VERSION : 0.1
   VAR
      ReadWriteDeviceNo : Int := 0;
      CopyDeviceNO : Int := 0;
      Read : Bool := FALSE;
      Write : Bool := FALSE;
      Copy : Bool := FALSE;
      Option : Array[0..2] of Struct
         With2PSwitch : Bool;
      END_STRUCT;
      MH_Hyd : Array[0..2] of "UDT721_Hydraulic";
      S_Hyd : Array[0..2] of "UDT721_Hydraulic";
      NZL_Hyd : Array[0..2] of "UDT721_Hydraulic";
   END_VAR
BEGIN
   MH_Hyd[0].Hyd_Filter_supervision := S5T#30S;
   MH_Hyd[0].Hyd_P_Startup := S5T#15S;
   MH_Hyd[0].Hyd_P_Supervision := S5T#5S;
   MH_Hyd[0].Hyd_CP_Time := S5T#4S;
   MH_Hyd[0].Hyd_PressureSwitch := S5T#0MS;
   MH_Hyd[0].Hyd_SwitchOFFDelay := S5T#0MS;
   MH_Hyd[1].Hyd_Filter_supervision := S5T#30S;
   MH_Hyd[1].Hyd_P_Startup := S5T#15S;
   MH_Hyd[1].Hyd_P_Supervision := S5T#5S;
   MH_Hyd[1].Hyd_CP_Time := S5T#4S;
   MH_Hyd[1].Hyd_PressureSwitch := S5T#0MS;
   MH_Hyd[1].Hyd_SwitchOFFDelay := S5T#0MS;
   MH_Hyd[2].Hyd_Filter_supervision := S5T#0MS;
   MH_Hyd[2].Hyd_P_Startup := S5T#0MS;
   MH_Hyd[2].Hyd_P_Supervision := S5T#0MS;
   MH_Hyd[2].Hyd_CP_Time := S5T#0MS;
   MH_Hyd[2].Hyd_PressureSwitch := S5T#0MS;
   MH_Hyd[2].Hyd_SwitchOFFDelay := S5T#0MS;
   S_Hyd[0].Hyd_Filter_supervision := S5T#0MS;
   S_Hyd[0].Hyd_P_Startup := S5T#0MS;
   S_Hyd[0].Hyd_P_Supervision := S5T#0MS;
   S_Hyd[0].Hyd_CP_Time := S5T#0MS;
   S_Hyd[0].Hyd_PressureSwitch := S5T#0MS;
   S_Hyd[0].Hyd_SwitchOFFDelay := S5T#0MS;
   S_Hyd[1].Hyd_Filter_supervision := S5T#0MS;
   S_Hyd[1].Hyd_P_Startup := S5T#0MS;
   S_Hyd[1].Hyd_P_Supervision := S5T#0MS;
   S_Hyd[1].Hyd_CP_Time := S5T#0MS;
   S_Hyd[1].Hyd_PressureSwitch := S5T#0MS;
   S_Hyd[1].Hyd_SwitchOFFDelay := S5T#0MS;
   S_Hyd[2].Hyd_Filter_supervision := S5T#0MS;
   S_Hyd[2].Hyd_P_Startup := S5T#0MS;
   S_Hyd[2].Hyd_P_Supervision := S5T#0MS;
   S_Hyd[2].Hyd_CP_Time := S5T#0MS;
   S_Hyd[2].Hyd_PressureSwitch := S5T#0MS;
   S_Hyd[2].Hyd_SwitchOFFDelay := S5T#0MS;
   NZL_Hyd[0].Hyd_Filter_supervision := S5T#0MS;
   NZL_Hyd[0].Hyd_P_Startup := S5T#0MS;
   NZL_Hyd[0].Hyd_P_Supervision := S5T#0MS;
   NZL_Hyd[0].Hyd_CP_Time := S5T#0MS;
   NZL_Hyd[0].Hyd_PressureSwitch := S5T#0MS;
   NZL_Hyd[0].Hyd_SwitchOFFDelay := S5T#0MS;
   NZL_Hyd[1].Hyd_Filter_supervision := S5T#0MS;
   NZL_Hyd[1].Hyd_P_Startup := S5T#0MS;
   NZL_Hyd[1].Hyd_P_Supervision := S5T#0MS;
   NZL_Hyd[1].Hyd_CP_Time := S5T#0MS;
   NZL_Hyd[1].Hyd_PressureSwitch := S5T#0MS;
   NZL_Hyd[1].Hyd_SwitchOFFDelay := S5T#0MS;
   NZL_Hyd[2].Hyd_Filter_supervision := S5T#0MS;
   NZL_Hyd[2].Hyd_P_Startup := S5T#0MS;
   NZL_Hyd[2].Hyd_P_Supervision := S5T#0MS;
   NZL_Hyd[2].Hyd_CP_Time := S5T#0MS;
   NZL_Hyd[2].Hyd_PressureSwitch := S5T#0MS;
   NZL_Hyd[2].Hyd_SwitchOFFDelay := S5T#0MS;
   Option[0].With2PSwitch := TRUE;
   Option[1].With2PSwitch := TRUE;
   Option[2].With2PSwitch := FALSE;
END_DATA_BLOCK

DATA_BLOCK "DB753_MeteringPump"   // DB753
TITLE = Parameter metering pump
{ S7_Optimized_Access := 'FALSE' }
NAME : metering
VERSION : 0.1
   VAR
      ReadWriteDeviceNo : Int := 0;
      CopyDeviceNO : Int := 0;
      Read : Bool := FALSE;
      Write : Bool := FALSE;
      Copy : Bool := FALSE;
      Pump : Array[0..12] of "UDT753_MeteringPump";
      Heating : Array[0..12] of Struct
         Exist : Array[1..8] of Bool;
      END_STRUCT;
      HeatingController : Array[0..4] of Struct
         Heating : Array[1..8] of "UDT702_HeatingControl";
      END_STRUCT;
   END_VAR
BEGIN
   Pump[0].Pump_Active := TRUE;
   Pump[0].WithFC := TRUE;
   Pump[0].WithoutFlowControl := TRUE;
   Pump[0].WithFeedPump := FALSE;
   Pump[0].WithEdgeFilter := FALSE;
   Pump[0].MachineNumber := 16#01;
   Pump[0]."Name" := 'Poly';
   Pump[0].TankNo := 1;
   Pump[0].Pulse_per_liter := 333.333;
   Pump[1].Pump_Active := TRUE;
   Pump[1].WithFC := TRUE;
   Pump[1].WithoutFlowControl := TRUE;
   Pump[1].WithFeedPump := FALSE;
   Pump[1].WithEdgeFilter := FALSE;
   Pump[1]."Name" := 'Poly';
   Pump[1].TankNo := 1;
   Pump[2].Pump_Active := TRUE;
   Pump[2].WithFC := TRUE;
   Pump[2].WithoutFlowControl := TRUE;
   Pump[2].WithFeedPump := FALSE;
   Pump[2].WithEdgeFilter := FALSE;
   Pump[2].MachineNumber := 16#01;
   Pump[2]."Name" := 'Iso';
   Pump[2].TankNo := 2;
   Pump[2].Pulse_per_liter := 965.667;
   Pump[0].Flow_State := 16#0000;
   Pump[0].RunTimePumpInterval := S5T#0MS;
   Pump[0].PauseTimePumpInterval := S5T#0MS;
   Pump[0].Flow_Index := 16#0000;
   Pump[0].DelayPressureFeedP := S5T#9S;
   Pump[0].DelayRunTimeFeedP := S5T#6S;
   Pump[0].MinTempRelease := 0.0;
   Pump[0].With_2Point := FALSE;
   Pump[0].WithFlowControl := FALSE;
   Pump[0].PumDeselectionEnable := FALSE;
   Pump[0].PumpDeselected := FALSE;
   Pump[0].PumpDeselectedInterval := FALSE;
   Pump[0].WithFischerValveHP := FALSE;
   Pump[0].WithFischerValveLP := FALSE;
   Pump[0].WithHPHeatExchanger := FALSE;
   Pump[0].WithLPHeatExchanger := FALSE;
   Pump[0].WithExhauseSystem := FALSE;
   Pump[0].WithHeating := FALSE;
   Pump[0].WithPipeHeating := FALSE;
   Pump[0].WithMinTempRelease := FALSE;
   Pump[0].WithFlowFactor := FALSE;
   Pump[0].With_1Speed := FALSE;
   Pump[0].With_2Speed := FALSE;
   Pump[0].WithExternalFan := FALSE;
   Pump[0].Spare23 := FALSE;
   Pump[0].Spare24 := FALSE;
   Pump[0].MaxFlowPercent := 100.0;
   Pump[0].MinFlowPercent := 10.0;
   Pump[0].MaxFlowLiter := 40.0;
   Pump[0].FlowFactor := 1.0;
   Pump[1].Flow_State := 16#0000;
   Pump[1].RunTimePumpInterval := S5T#0MS;
   Pump[1].PauseTimePumpInterval := S5T#0MS;
   Pump[1].Flow_Index := 16#0000;
   Pump[1].DelayPressureFeedP := S5T#9S;
   Pump[1].DelayRunTimeFeedP := S5T#6S;
   Pump[1].MinTempRelease := 0.0;
   Pump[1].With_2Point := FALSE;
   Pump[1].WithFlowControl := FALSE;
   Pump[1].PumDeselectionEnable := FALSE;
   Pump[1].PumpDeselected := FALSE;
   Pump[1].PumpDeselectedInterval := FALSE;
   Pump[1].WithFischerValveHP := FALSE;
   Pump[1].WithFischerValveLP := FALSE;
   Pump[1].WithHPHeatExchanger := FALSE;
   Pump[1].WithLPHeatExchanger := FALSE;
   Pump[1].WithExhauseSystem := FALSE;
   Pump[1].WithHeating := FALSE;
   Pump[1].WithPipeHeating := FALSE;
   Pump[1].WithMinTempRelease := FALSE;
   Pump[1].WithFlowFactor := FALSE;
   Pump[1].With_1Speed := FALSE;
   Pump[1].With_2Speed := FALSE;
   Pump[1].WithExternalFan := FALSE;
   Pump[1].Spare23 := FALSE;
   Pump[1].Spare24 := FALSE;
   Pump[1].MachineNumber := 16#01;
   Pump[1].Pulse_per_liter := 333.333;
   Pump[1].MaxFlowPercent := 100.0;
   Pump[1].MinFlowPercent := 10.0;
   Pump[1].MaxFlowLiter := 40.0;
   Pump[1].FlowFactor := 1.0;
   Pump[2].Flow_State := 16#0000;
   Pump[2].RunTimePumpInterval := S5T#0MS;
   Pump[2].PauseTimePumpInterval := S5T#0MS;
   Pump[2].Flow_Index := 16#0000;
   Pump[2].DelayPressureFeedP := S5T#10S;
   Pump[2].DelayRunTimeFeedP := S5T#5S;
   Pump[2].MinTempRelease := 0.0;
   Pump[2].With_2Point := FALSE;
   Pump[2].WithFlowControl := FALSE;
   Pump[2].PumDeselectionEnable := FALSE;
   Pump[2].PumpDeselected := FALSE;
   Pump[2].PumpDeselectedInterval := FALSE;
   Pump[2].WithFischerValveHP := FALSE;
   Pump[2].WithFischerValveLP := FALSE;
   Pump[2].WithHPHeatExchanger := FALSE;
   Pump[2].WithLPHeatExchanger := FALSE;
   Pump[2].WithExhauseSystem := FALSE;
   Pump[2].WithHeating := FALSE;
   Pump[2].WithPipeHeating := FALSE;
   Pump[2].WithMinTempRelease := FALSE;
   Pump[2].WithFlowFactor := FALSE;
   Pump[2].With_1Speed := FALSE;
   Pump[2].With_2Speed := FALSE;
   Pump[2].WithExternalFan := FALSE;
   Pump[2].Spare23 := FALSE;
   Pump[2].Spare24 := FALSE;
   Pump[2].MaxFlowPercent := 100.0;
   Pump[2].MinFlowPercent := 10.0;
   Pump[2].MaxFlowLiter := 16.0;
   Pump[2].FlowFactor := 1.0;
   Pump[3].Flow_State := 16#0000;
   Pump[3].RunTimePumpInterval := S5T#0MS;
   Pump[3].PauseTimePumpInterval := S5T#0MS;
   Pump[3].Flow_Index := 16#0000;
   Pump[3].DelayPressureFeedP := S5T#0MS;
   Pump[3].DelayRunTimeFeedP := S5T#0MS;
   Pump[3].MinTempRelease := 0.0;
   Pump[3].Pump_Active := FALSE;
   Pump[3].WithFC := FALSE;
   Pump[3].With_2Point := FALSE;
   Pump[3].WithFlowControl := FALSE;
   Pump[3].WithoutFlowControl := FALSE;
   Pump[3].WithFeedPump := FALSE;
   Pump[3].WithEdgeFilter := FALSE;
   Pump[3].PumDeselectionEnable := FALSE;
   Pump[3].PumpDeselected := FALSE;
   Pump[3].PumpDeselectedInterval := FALSE;
   Pump[3].WithFischerValveHP := FALSE;
   Pump[3].WithFischerValveLP := FALSE;
   Pump[3].WithHPHeatExchanger := FALSE;
   Pump[3].WithLPHeatExchanger := FALSE;
   Pump[3].WithExhauseSystem := FALSE;
   Pump[3].WithHeating := FALSE;
   Pump[3].WithPipeHeating := FALSE;
   Pump[3].WithMinTempRelease := FALSE;
   Pump[3].WithFlowFactor := FALSE;
   Pump[3].With_1Speed := FALSE;
   Pump[3].With_2Speed := FALSE;
   Pump[3].WithExternalFan := FALSE;
   Pump[3].Spare23 := FALSE;
   Pump[3].Spare24 := FALSE;
   Pump[3].MachineNumber := 16#01;
   Pump[3]."Name" := 'Comp 03';
   Pump[3].TankNo := 3;
   Pump[3].Pulse_per_liter := 965.0;
   Pump[3].MaxFlowPercent := 0.0;
   Pump[3].MinFlowPercent := 0.0;
   Pump[3].MaxFlowLiter := 0.0;
   Pump[3].FlowFactor := 0.0;
   Pump[4].Flow_State := 16#0000;
   Pump[4].RunTimePumpInterval := S5T#0MS;
   Pump[4].PauseTimePumpInterval := S5T#0MS;
   Pump[4].Flow_Index := 16#0000;
   Pump[4].DelayPressureFeedP := S5T#0MS;
   Pump[4].DelayRunTimeFeedP := S5T#0MS;
   Pump[4].MinTempRelease := 0.0;
   Pump[4].Pump_Active := FALSE;
   Pump[4].WithFC := FALSE;
   Pump[4].With_2Point := FALSE;
   Pump[4].WithFlowControl := FALSE;
   Pump[4].WithoutFlowControl := FALSE;
   Pump[4].WithFeedPump := FALSE;
   Pump[4].WithEdgeFilter := FALSE;
   Pump[4].PumDeselectionEnable := FALSE;
   Pump[4].PumpDeselected := FALSE;
   Pump[4].PumpDeselectedInterval := FALSE;
   Pump[4].WithFischerValveHP := FALSE;
   Pump[4].WithFischerValveLP := FALSE;
   Pump[4].WithHPHeatExchanger := FALSE;
   Pump[4].WithLPHeatExchanger := FALSE;
   Pump[4].WithExhauseSystem := FALSE;
   Pump[4].WithHeating := FALSE;
   Pump[4].WithPipeHeating := FALSE;
   Pump[4].WithMinTempRelease := FALSE;
   Pump[4].WithFlowFactor := FALSE;
   Pump[4].With_1Speed := FALSE;
   Pump[4].With_2Speed := FALSE;
   Pump[4].WithExternalFan := FALSE;
   Pump[4].Spare23 := FALSE;
   Pump[4].Spare24 := FALSE;
   Pump[4].MachineNumber := 16#01;
   Pump[4]."Name" := 'Comp 04';
   Pump[4].TankNo := 4;
   Pump[4].Pulse_per_liter := 965.0;
   Pump[4].MaxFlowLiter := 0.0;
   Pump[4].MinFlowPercent := 0.0;
   Pump[4].MaxFlowPercent := 0.0;
   Pump[4].FlowFactor := 0.0;
   Pump[5].Flow_State := 16#0000;
   Pump[5].RunTimePumpInterval := S5T#0MS;
   Pump[5].PauseTimePumpInterval := S5T#0MS;
   Pump[5].Flow_Index := 16#0000;
   Pump[5].DelayPressureFeedP := S5T#0MS;
   // 557 more start values not shown
END_DATA_BLOCK

DATA_BLOCK "DB761_Cylinder_Manager"   // DB761
TITLE = Parameter cylinder manager
{ S7_Optimized_Access := 'FALSE' }
VERSION : 0.1
   VAR
      ReadWriteDeviceNo : Int := 0;
      CopyDeviceNO : Int := 0;
      Read : Bool := FALSE;
      Write : Bool := FALSE;
      Copy : Bool := FALSE;
      CylinderMan_Ma : Array[0..2] of "UDT761_CylinderManager";
   END_VAR
BEGIN
   CylinderMan_Ma[0].Preparation_Cylinder := S5T#0MS;
   CylinderMan_Ma[0].PausePos_Auto := 0;
   CylinderMan_Ma[0].PausePos_Manual := 0;
   CylinderMan_Ma[0].reserve_01 := 0;
   CylinderMan_Ma[0].reserve_02 := 0;
   CylinderMan_Ma[0].reserve_03 := 0;
   CylinderMan_Ma[1].Preparation_Cylinder := S5T#0MS;
   CylinderMan_Ma[1].PausePos_Auto := 0;
   CylinderMan_Ma[1].PausePos_Manual := 0;
   CylinderMan_Ma[1].reserve_01 := 0;
   CylinderMan_Ma[1].reserve_02 := 0;
   CylinderMan_Ma[1].reserve_03 := 0;
   CylinderMan_Ma[2].Preparation_Cylinder := S5T#0MS;
   CylinderMan_Ma[2].PausePos_Auto := 0;
   CylinderMan_Ma[2].PausePos_Manual := 0;
   CylinderMan_Ma[2].reserve_01 := 0;
   CylinderMan_Ma[2].reserve_02 := 0;
   CylinderMan_Ma[2].reserve_03 := 0;
END_DATA_BLOCK

DATA_BLOCK "DB762_Cylinder"   // DB762
TITLE = Parameter cylinder
{ S7_Optimized_Access := 'FALSE' }
VERSION : 0.1
   VAR
      ReadWriteDeviceNo : Int := 0;
      CopyDeviceNO : Int := 0;
      Read : Bool := FALSE;
      Write : Bool := FALSE;
      Copy : Bool := FALSE;
      Cylinder : Array[0..12] of "UDT762_Cylinder";
   END_VAR
BEGIN
   Cylinder[0].Cyl_PausePosition_Auto := FALSE;
   Cylinder[0].Cyl_PausePosition_Manual := FALSE;
   Cylinder[0].Spare_02 := FALSE;
   Cylinder[0].Spare_03 := FALSE;
   Cylinder[0].Spare_04 := FALSE;
   Cylinder[0].Spare_05 := FALSE;
   Cylinder[0].Spare_06 := FALSE;
   Cylinder[0].Spare_07 := FALSE;
   Cylinder[0].No_cyl_cycle_lubricate := 0;
   Cylinder[0].Spare_6 := 0;
   Cylinder[0].Spare_8 := 0;
   Cylinder[0].T_SetValMeterAfterValve := S5T#0MS;
   Cylinder[0].T_ValveMeterAfterSetVal := S5T#0MS;
   Cylinder[0].T_PistonVenting := S5T#0MS;
   Cylinder[0].T_PauseAfterMetering := S5T#0MS;
   Cylinder[0].T_FillValPreSuctionVal := S5T#0MS;
   Cylinder[0].T_SetValFillAfterValve := S5T#0MS;
   Cylinder[0].T_ValveFillAfterSetVal := S5T#0MS;
   Cylinder[0].T_PauseAfterFilling := S5T#0MS;
   Cylinder[0].T_MonitoringPBFeedpump := S5T#0MS;
   Cylinder[0].Spare26 := 0;
   Cylinder[0].SetValueFilling := 0;
   Cylinder[0].SetVMeteringCylSer := 0;
   Cylinder[0].SetVFillingCylSer := 0;
   Cylinder[1].Cyl_PausePosition_Auto := FALSE;
   Cylinder[1].Cyl_PausePosition_Manual := FALSE;
   Cylinder[1].Spare_02 := FALSE;
   Cylinder[1].Spare_03 := FALSE;
   Cylinder[1].Spare_04 := FALSE;
   Cylinder[1].Spare_05 := FALSE;
   Cylinder[1].Spare_06 := FALSE;
   Cylinder[1].Spare_07 := FALSE;
   Cylinder[1].No_cyl_cycle_lubricate := 0;
   Cylinder[1].Spare_6 := 0;
   Cylinder[1].Spare_8 := 0;
   Cylinder[1].T_SetValMeterAfterValve := S5T#0MS;
   Cylinder[1].T_ValveMeterAfterSetVal := S5T#0MS;
   Cylinder[1].T_PistonVenting := S5T#0MS;
   Cylinder[1].T_PauseAfterMetering := S5T#0MS;
   Cylinder[1].T_FillValPreSuctionVal := S5T#0MS;
   Cylinder[1].T_SetValFillAfterValve := S5T#0MS;
   Cylinder[1].T_ValveFillAfterSetVal := S5T#0MS;
   Cylinder[1].T_PauseAfterFilling := S5T#0MS;
   Cylinder[1].T_MonitoringPBFeedpump := S5T#0MS;
   Cylinder[1].Spare26 := 0;
   Cylinder[1].SetValueFilling := 0;
   Cylinder[1].SetVMeteringCylSer := 0;
   Cylinder[1].SetVFillingCylSer := 0;
   Cylinder[2].Cyl_PausePosition_Auto := FALSE;
   Cylinder[2].Cyl_PausePosition_Manual := FALSE;
   Cylinder[2].Spare_02 := FALSE;
   Cylinder[2].Spare_03 := FALSE;
   Cylinder[2].Spare_04 := FALSE;
   Cylinder[2].Spare_05 := FALSE;
   Cylinder[2].Spare_06 := FALSE;
   Cylinder[2].Spare_07 := FALSE;
   Cylinder[2].No_cyl_cycle_lubricate := 0;
   Cylinder[2].Spare_6 := 0;
   Cylinder[2].Spare_8 := 0;
   Cylinder[2].T_SetValMeterAfterValve := S5T#0MS;
   Cylinder[2].T_ValveMeterAfterSetVal := S5T#0MS;
   Cylinder[2].T_PistonVenting := S5T#0MS;
   Cylinder[2].T_PauseAfterMetering := S5T#0MS;
   Cylinder[2].T_FillValPreSuctionVal := S5T#0MS;
   Cylinder[2].T_SetValFillAfterValve := S5T#0MS;
   Cylinder[2].T_ValveFillAfterSetVal := S5T#0MS;
   Cylinder[2].T_PauseAfterFilling := S5T#0MS;
   Cylinder[2].T_MonitoringPBFeedpump := S5T#0MS;
   Cylinder[2].Spare26 := 0;
   Cylinder[2].SetValueFilling := 0;
   Cylinder[2].SetVMeteringCylSer := 0;
   Cylinder[2].SetVFillingCylSer := 0;
   Cylinder[3].Cyl_PausePosition_Auto := FALSE;
   Cylinder[3].Cyl_PausePosition_Manual := FALSE;
   Cylinder[3].Spare_02 := FALSE;
   Cylinder[3].Spare_03 := FALSE;
   Cylinder[3].Spare_04 := FALSE;
   Cylinder[3].Spare_05 := FALSE;
   Cylinder[3].Spare_06 := FALSE;
   Cylinder[3].Spare_07 := FALSE;
   Cylinder[3].No_cyl_cycle_lubricate := 0;
   Cylinder[3].Spare_6 := 0;
   Cylinder[3].Spare_8 := 0;
   Cylinder[3].T_SetValMeterAfterValve := S5T#0MS;
   Cylinder[3].T_ValveMeterAfterSetVal := S5T#0MS;
   Cylinder[3].T_PistonVenting := S5T#0MS;
   Cylinder[3].T_PauseAfterMetering := S5T#0MS;
   Cylinder[3].T_FillValPreSuctionVal := S5T#0MS;
   Cylinder[3].T_SetValFillAfterValve := S5T#0MS;
   Cylinder[3].T_ValveFillAfterSetVal := S5T#0MS;
   Cylinder[3].T_PauseAfterFilling := S5T#0MS;
   Cylinder[3].T_MonitoringPBFeedpump := S5T#0MS;
   Cylinder[3].Spare26 := 0;
   Cylinder[3].SetValueFilling := 0;
   Cylinder[3].SetVMeteringCylSer := 0;
   Cylinder[3].SetVFillingCylSer := 0;
   Cylinder[4].Cyl_PausePosition_Auto := FALSE;
   Cylinder[4].Cyl_PausePosition_Manual := FALSE;
   Cylinder[4].Spare_02 := FALSE;
   Cylinder[4].Spare_03 := FALSE;
   Cylinder[4].Spare_04 := FALSE;
   Cylinder[4].Spare_05 := FALSE;
   Cylinder[4].Spare_06 := FALSE;
   Cylinder[4].Spare_07 := FALSE;
   Cylinder[4].No_cyl_cycle_lubricate := 0;
   Cylinder[4].Spare_6 := 0;
   Cylinder[4].Spare_8 := 0;
   Cylinder[4].T_SetValMeterAfterValve := S5T#0MS;
   Cylinder[4].T_ValveMeterAfterSetVal := S5T#0MS;
   Cylinder[4].T_PistonVenting := S5T#0MS;
   Cylinder[4].T_PauseAfterMetering := S5T#0MS;
   Cylinder[4].T_FillValPreSuctionVal := S5T#0MS;
   Cylinder[4].T_SetValFillAfterValve := S5T#0MS;
   Cylinder[4].T_ValveFillAfterSetVal := S5T#0MS;
   Cylinder[4].T_PauseAfterFilling := S5T#0MS;
   Cylinder[4].T_MonitoringPBFeedpump := S5T#0MS;
   Cylinder[4].Spare26 := 0;
   Cylinder[4].SetValueFilling := 0;
   Cylinder[4].SetVMeteringCylSer := 0;
   Cylinder[4].SetVFillingCylSer := 0;
   Cylinder[5].Cyl_PausePosition_Auto := FALSE;
   Cylinder[5].Cyl_PausePosition_Manual := FALSE;
   Cylinder[5].Spare_02 := FALSE;
   Cylinder[5].Spare_03 := FALSE;
   Cylinder[5].Spare_04 := FALSE;
   Cylinder[5].Spare_05 := FALSE;
   Cylinder[5].Spare_06 := FALSE;
   Cylinder[5].Spare_07 := FALSE;
   Cylinder[5].No_cyl_cycle_lubricate := 0;
   Cylinder[5].Spare_6 := 0;
   Cylinder[5].Spare_8 := 0;
   Cylinder[5].T_SetValMeterAfterValve := S5T#0MS;
   Cylinder[5].T_ValveMeterAfterSetVal := S5T#0MS;
   Cylinder[5].T_PistonVenting := S5T#0MS;
   Cylinder[5].T_PauseAfterMetering := S5T#0MS;
   Cylinder[5].T_FillValPreSuctionVal := S5T#0MS;
   Cylinder[5].T_SetValFillAfterValve := S5T#0MS;
   Cylinder[5].T_ValveFillAfterSetVal := S5T#0MS;
   Cylinder[5].T_PauseAfterFilling := S5T#0MS;
   Cylinder[5].T_MonitoringPBFeedpump := S5T#0MS;
   Cylinder[5].Spare26 := 0;
   Cylinder[5].SetValueFilling := 0;
   Cylinder[5].SetVMeteringCylSer := 0;
   Cylinder[5].SetVFillingCylSer := 0;
   Cylinder[6].Cyl_PausePosition_Auto := FALSE;
   Cylinder[6].Cyl_PausePosition_Manual := FALSE;
   Cylinder[6].Spare_02 := FALSE;
   Cylinder[6].Spare_03 := FALSE;
   Cylinder[6].Spare_04 := FALSE;
   Cylinder[6].Spare_05 := FALSE;
   Cylinder[6].Spare_06 := FALSE;
   Cylinder[6].Spare_07 := FALSE;
   Cylinder[6].No_cyl_cycle_lubricate := 0;
   Cylinder[6].Spare_6 := 0;
   Cylinder[6].Spare_8 := 0;
   Cylinder[6].T_SetValMeterAfterValve := S5T#0MS;
   Cylinder[6].T_ValveMeterAfterSetVal := S5T#0MS;
   Cylinder[6].T_PistonVenting := S5T#0MS;
   Cylinder[6].T_PauseAfterMetering := S5T#0MS;
   Cylinder[6].T_FillValPreSuctionVal := S5T#0MS;
   Cylinder[6].T_SetValFillAfterValve := S5T#0MS;
   Cylinder[6].T_ValveFillAfterSetVal := S5T#0MS;
   Cylinder[6].T_PauseAfterFilling := S5T#0MS;
   Cylinder[6].T_MonitoringPBFeedpump := S5T#0MS;
   Cylinder[6].Spare26 := 0;
   Cylinder[6].SetValueFilling := 0;
   Cylinder[6].SetVMeteringCylSer := 0;
   Cylinder[6].SetVFillingCylSer := 0;
   Cylinder[7].Cyl_PausePosition_Auto := FALSE;
   Cylinder[7].Cyl_PausePosition_Manual := FALSE;
   Cylinder[7].Spare_02 := FALSE;
   Cylinder[7].Spare_03 := FALSE;
   Cylinder[7].Spare_04 := FALSE;
   Cylinder[7].Spare_05 := FALSE;
   Cylinder[7].Spare_06 := FALSE;
   Cylinder[7].Spare_07 := FALSE;
   Cylinder[7].No_cyl_cycle_lubricate := 0;
   Cylinder[7].Spare_6 := 0;
   Cylinder[7].Spare_8 := 0;
   Cylinder[7].T_SetValMeterAfterValve := S5T#0MS;
   Cylinder[7].T_ValveMeterAfterSetVal := S5T#0MS;
   Cylinder[7].T_PistonVenting := S5T#0MS;
   Cylinder[7].T_PauseAfterMetering := S5T#0MS;
   Cylinder[7].T_FillValPreSuctionVal := S5T#0MS;
   Cylinder[7].T_SetValFillAfterValve := S5T#0MS;
   Cylinder[7].T_ValveFillAfterSetVal := S5T#0MS;
   Cylinder[7].T_PauseAfterFilling := S5T#0MS;
   Cylinder[7].T_MonitoringPBFeedpump := S5T#0MS;
   Cylinder[7].Spare26 := 0;
   Cylinder[7].SetValueFilling := 0;
   Cylinder[7].SetVMeteringCylSer := 0;
   Cylinder[7].SetVFillingCylSer := 0;
   Cylinder[8].Cyl_PausePosition_Auto := FALSE;
   Cylinder[8].Cyl_PausePosition_Manual := FALSE;
   Cylinder[8].Spare_02 := FALSE;
   Cylinder[8].Spare_03 := FALSE;
   Cylinder[8].Spare_04 := FALSE;
   Cylinder[8].Spare_05 := FALSE;
   Cylinder[8].Spare_06 := FALSE;
   Cylinder[8].Spare_07 := FALSE;
   // 112 more start values not shown
END_DATA_BLOCK

DATA_BLOCK "DB790_PlantParameter"   // DB790
TITLE = Parameter plant
{ S7_Optimized_Access := 'FALSE' }
VERSION : 0.1
   VAR
      Bit : Struct
         WithRobots : Bool := FALSE;
         withTT : Bool := FALSE;
         MHNofromInterface : Bool := FALSE;   // Mixinghead No comes from Interface No
         ProgrammNofromInterface : Bool;   // Programm number comes from the interface
      END_STRUCT;
      AmountProCanModul : Int := 2;
      AmountMH : Int := 1;
      AmountTank : Int := 2;
      AmountMeteringUnits : Int := 2;
      AmountToolStation : Int := 1;   // Amount tools at a station
      AmountMouldCarrier : Int := 0;   // Amount mouldcarrier at a plant
      TestProgPerMH : Int := 99;   // Number of test programs per mixing head
      AmountToolAllocations : Int := 128;   // Amount of program numbers to start a foaming cycle
      MaxAmountShotAtTool : Int := 8;
      AmountRecipes : Int := 99;   // Amount of recipes at a plant
      AmountShots : Int := 255;   // Amount of shots at a plant
      AmountMachine : Int := 1;   // Amount machine at a plant
      AmountRobots : Int := 0;   // Amount robots at a plant
   END_VAR
BEGIN
END_DATA_BLOCK

DATA_BLOCK "DB820_Error_general"   // DB820
TITLE = Faults general at plant and machine
{ S7_Optimized_Access := 'FALSE' }
VERSION : 0.1
   VAR
      Profibus_DP : Array[0..2] of "UDT1805_FLT_PB_DP";   // Fault DP-member 1-10 fault level 1 others fault level 3
      Machine : Array[0..2] of "UDT1800_FLT_Machine";   // Machine general faults
   END_VAR
BEGIN
   Profibus_DP[0].Member[1] := FALSE;
   Profibus_DP[0].Member[2] := FALSE;
   Profibus_DP[0].Member[3] := FALSE;
   Profibus_DP[0].Member[4] := FALSE;
   Profibus_DP[0].Member[5] := FALSE;
   Profibus_DP[0].Member[6] := FALSE;
   Profibus_DP[0].Member[7] := FALSE;
   Profibus_DP[0].Member[8] := FALSE;
   Profibus_DP[0].Member[9] := FALSE;
   Profibus_DP[0].Member[10] := FALSE;
   Profibus_DP[0].Member[11] := FALSE;
   Profibus_DP[0].Member[12] := FALSE;
   Profibus_DP[0].Member[13] := FALSE;
   Profibus_DP[0].Member[14] := FALSE;
   Profibus_DP[0].Member[15] := FALSE;
   Profibus_DP[0].Member[16] := FALSE;
   Profibus_DP[0].Member[17] := FALSE;
   Profibus_DP[0].Member[18] := FALSE;
   Profibus_DP[0].Member[19] := FALSE;
   Profibus_DP[0].Member[20] := FALSE;
   Profibus_DP[0].Member[21] := FALSE;
   Profibus_DP[0].Member[22] := FALSE;
   Profibus_DP[0].Member[23] := FALSE;
   Profibus_DP[0].Member[24] := FALSE;
   Profibus_DP[0].Member[25] := FALSE;
   Profibus_DP[0].Member[26] := FALSE;
   Profibus_DP[0].Member[27] := FALSE;
   Profibus_DP[0].Member[28] := FALSE;
   Profibus_DP[0].Member[29] := FALSE;
   Profibus_DP[0].Member[30] := FALSE;
   Profibus_DP[0].Member[31] := FALSE;
   Profibus_DP[0].Member[32] := FALSE;
   Profibus_DP[0].Member[33] := FALSE;
   Profibus_DP[0].Member[34] := FALSE;
   Profibus_DP[0].Member[35] := FALSE;
   Profibus_DP[0].Member[36] := FALSE;
   Profibus_DP[0].Member[37] := FALSE;
   Profibus_DP[0].Member[38] := FALSE;
   Profibus_DP[0].Member[39] := FALSE;
   Profibus_DP[0].Member[40] := FALSE;
   Profibus_DP[0].Member[41] := FALSE;
   Profibus_DP[0].Member[42] := FALSE;
   Profibus_DP[0].Member[43] := FALSE;
   Profibus_DP[0].Member[44] := FALSE;
   Profibus_DP[0].Member[45] := FALSE;
   Profibus_DP[0].Member[46] := FALSE;
   Profibus_DP[0].Member[47] := FALSE;
   Profibus_DP[0].Member[48] := FALSE;
   Profibus_DP[0].Member[49] := FALSE;
   Profibus_DP[0].Member[50] := FALSE;
   Profibus_DP[0].Member[51] := FALSE;
   Profibus_DP[0].Member[52] := FALSE;
   Profibus_DP[0].Member[53] := FALSE;
   Profibus_DP[0].Member[54] := FALSE;
   Profibus_DP[0].Member[55] := FALSE;
   Profibus_DP[0].Member[56] := FALSE;
   Profibus_DP[0].Member[57] := FALSE;
   Profibus_DP[0].Member[58] := FALSE;
   Profibus_DP[0].Member[59] := FALSE;
   Profibus_DP[0].Member[60] := FALSE;
   Profibus_DP[0].Member[61] := FALSE;
   Profibus_DP[0].Member[62] := FALSE;
   Profibus_DP[0].Member[63] := FALSE;
   Profibus_DP[0].Member[64] := FALSE;
   Profibus_DP[0].Member[65] := FALSE;
   Profibus_DP[0].Member[66] := FALSE;
   Profibus_DP[0].Member[67] := FALSE;
   Profibus_DP[0].Member[68] := FALSE;
   Profibus_DP[0].Member[69] := FALSE;
   Profibus_DP[0].Member[70] := FALSE;
   Profibus_DP[0].Member[71] := FALSE;
   Profibus_DP[0].Member[72] := FALSE;
   Profibus_DP[0].Member[73] := FALSE;
   Profibus_DP[0].Member[74] := FALSE;
   Profibus_DP[0].Member[75] := FALSE;
   Profibus_DP[0].Member[76] := FALSE;
   Profibus_DP[0].Member[77] := FALSE;
   Profibus_DP[0].Member[78] := FALSE;
   Profibus_DP[0].Member[79] := FALSE;
   Profibus_DP[0].Member[80] := FALSE;
   Profibus_DP[0].Member[81] := FALSE;
   Profibus_DP[0].Member[82] := FALSE;
   Profibus_DP[0].Member[83] := FALSE;
   Profibus_DP[0].Member[84] := FALSE;
   Profibus_DP[0].Member[85] := FALSE;
   Profibus_DP[0].Member[86] := FALSE;
   Profibus_DP[0].Member[87] := FALSE;
   Profibus_DP[0].Member[88] := FALSE;
   Profibus_DP[0].Member[89] := FALSE;
   Profibus_DP[0].Member[90] := FALSE;
   Profibus_DP[0].Member[91] := FALSE;
   Profibus_DP[0].Member[92] := FALSE;
   Profibus_DP[0].Member[93] := FALSE;
   Profibus_DP[0].Member[94] := FALSE;
   Profibus_DP[0].Member[95] := FALSE;
   Profibus_DP[0].Member[96] := FALSE;
   Profibus_DP[0].Member[97] := FALSE;
   Profibus_DP[0].Member[98] := FALSE;
   Profibus_DP[0].Member[99] := FALSE;
   Profibus_DP[0].Member[100] := FALSE;
   Profibus_DP[0].Member[101] := FALSE;
   Profibus_DP[0].Member[102] := FALSE;
   Profibus_DP[0].Member[103] := FALSE;
   Profibus_DP[0].Member[104] := FALSE;
   Profibus_DP[0].Member[105] := FALSE;
   Profibus_DP[0].Member[106] := FALSE;
   Profibus_DP[0].Member[107] := FALSE;
   Profibus_DP[0].Member[108] := FALSE;
   Profibus_DP[0].Member[109] := FALSE;
   Profibus_DP[0].Member[110] := FALSE;
   Profibus_DP[0].Member[111] := FALSE;
   Profibus_DP[0].Member[112] := FALSE;
   Profibus_DP[0].Member[113] := FALSE;
   Profibus_DP[0].Member[114] := FALSE;
   Profibus_DP[0].Member[115] := FALSE;
   Profibus_DP[0].Member[116] := FALSE;
   Profibus_DP[0].Member[117] := FALSE;
   Profibus_DP[0].Member[118] := FALSE;
   Profibus_DP[0].Member[119] := FALSE;
   Profibus_DP[0].Member[120] := FALSE;
   Profibus_DP[0].Member[121] := FALSE;
   Profibus_DP[0].Member[122] := FALSE;
   Profibus_DP[0].Member[123] := FALSE;
   Profibus_DP[0].Member[124] := FALSE;
   Profibus_DP[0].Member[125] := FALSE;
   Profibus_DP[0].Member[126] := FALSE;
   Profibus_DP[0].Member[127] := FALSE;
   Profibus_DP[0].Member[128] := FALSE;
   Profibus_DP[1].Member[1] := FALSE;
   Profibus_DP[1].Member[2] := FALSE;
   Profibus_DP[1].Member[3] := FALSE;
   Profibus_DP[1].Member[4] := FALSE;
   Profibus_DP[1].Member[5] := FALSE;
   Profibus_DP[1].Member[6] := FALSE;
   Profibus_DP[1].Member[7] := FALSE;
   Profibus_DP[1].Member[8] := FALSE;
   Profibus_DP[1].Member[9] := FALSE;
   Profibus_DP[1].Member[10] := FALSE;
   Profibus_DP[1].Member[11] := FALSE;
   Profibus_DP[1].Member[12] := FALSE;
   Profibus_DP[1].Member[13] := FALSE;
   Profibus_DP[1].Member[14] := FALSE;
   Profibus_DP[1].Member[15] := FALSE;
   Profibus_DP[1].Member[16] := FALSE;
   Profibus_DP[1].Member[17] := FALSE;
   Profibus_DP[1].Member[18] := FALSE;
   Profibus_DP[1].Member[19] := FALSE;
   Profibus_DP[1].Member[20] := FALSE;
   Profibus_DP[1].Member[21] := FALSE;
   Profibus_DP[1].Member[22] := FALSE;
   Profibus_DP[1].Member[23] := FALSE;
   Profibus_DP[1].Member[24] := FALSE;
   Profibus_DP[1].Member[25] := FALSE;
   Profibus_DP[1].Member[26] := FALSE;
   Profibus_DP[1].Member[27] := FALSE;
   Profibus_DP[1].Member[28] := FALSE;
   Profibus_DP[1].Member[29] := FALSE;
   Profibus_DP[1].Member[30] := FALSE;
   Profibus_DP[1].Member[31] := FALSE;
   Profibus_DP[1].Member[32] := FALSE;
   Profibus_DP[1].Member[33] := FALSE;
   Profibus_DP[1].Member[34] := FALSE;
   Profibus_DP[1].Member[35] := FALSE;
   Profibus_DP[1].Member[36] := FALSE;
   Profibus_DP[1].Member[37] := FALSE;
   Profibus_DP[1].Member[38] := FALSE;
   Profibus_DP[1].Member[39] := FALSE;
   Profibus_DP[1].Member[40] := FALSE;
   Profibus_DP[1].Member[41] := FALSE;
   Profibus_DP[1].Member[42] := FALSE;
   Profibus_DP[1].Member[43] := FALSE;
   Profibus_DP[1].Member[44] := FALSE;
   Profibus_DP[1].Member[45] := FALSE;
   Profibus_DP[1].Member[46] := FALSE;
   Profibus_DP[1].Member[47] := FALSE;
   Profibus_DP[1].Member[48] := FALSE;
   Profibus_DP[1].Member[49] := FALSE;
   Profibus_DP[1].Member[50] := FALSE;
   Profibus_DP[1].Member[51] := FALSE;
   Profibus_DP[1].Member[52] := FALSE;
   Profibus_DP[1].Member[53] := FALSE;
   Profibus_DP[1].Member[54] := FALSE;
   Profibus_DP[1].Member[55] := FALSE;
   Profibus_DP[1].Member[56] := FALSE;
   Profibus_DP[1].Member[57] := FALSE;
   Profibus_DP[1].Member[58] := FALSE;
   Profibus_DP[1].Member[59] := FALSE;
   Profibus_DP[1].Member[60] := FALSE;
   Profibus_DP[1].Member[61] := FALSE;
   Profibus_DP[1].Member[62] := FALSE;
   Profibus_DP[1].Member[63] := FALSE;
   Profibus_DP[1].Member[64] := FALSE;
   Profibus_DP[1].Member[65] := FALSE;
   Profibus_DP[1].Member[66] := FALSE;
   Profibus_DP[1].Member[67] := FALSE;
   Profibus_DP[1].Member[68] := FALSE;
   Profibus_DP[1].Member[69] := FALSE;
   Profibus_DP[1].Member[70] := FALSE;
   Profibus_DP[1].Member[71] := FALSE;
   Profibus_DP[1].Member[72] := FALSE;
   // 424 more start values not shown
END_DATA_BLOCK

DATA_BLOCK "DB821_Error_Hydraulic"   // DB821
TITLE = Faults general at plant and machine
{ S7_Optimized_Access := 'FALSE' }
VERSION : 0.1
   VAR
      MH_Hydraulic : Array[0..2] of "UDT1821_FLT_MH_Hydraulic";   // Mixinghead hydraulic
      S_Hydraulic : Array[0..2] of "UDT1821_FLT_MH_Hydraulic";   // Servo hydraulic
      NZL_Hydraulic : Array[0..2] of "UDT1821_FLT_MH_Hydraulic";   // Nozzle hydraulic
      EmergencyStop_Hydraulic : Array[1..16] of Bool;
   END_VAR
BEGIN
   MH_Hydraulic[0].FLT_Motorprotection := FALSE;
   MH_Hydraulic[0].FLT_Min_Level := FALSE;
   MH_Hydraulic[0].FLT_WRN_C_Max := FALSE;
   MH_Hydraulic[0].FLT_C_Max := FALSE;
   MH_Hydraulic[0].FLT_Filter_HP := FALSE;
   MH_Hydraulic[0].FLT_Filter_backflow := FALSE;
   MH_Hydraulic[0].FLT_cable_break := FALSE;
   MH_Hydraulic[0].FLT_P_Max := FALSE;
   MH_Hydraulic[0].FLT_Moog_Filter := FALSE;
   MH_Hydraulic[0].FLT_MotorProtFilterPump := FALSE;
   MH_Hydraulic[0].FLT_MinLevelFilterPump := FALSE;
   MH_Hydraulic[0].FLT_MaxLevelFilterPump := FALSE;
   MH_Hydraulic[0].FLT_FilterBypass := FALSE;
   MH_Hydraulic[0].Spare14 := FALSE;
   MH_Hydraulic[0].Spare15 := FALSE;
   MH_Hydraulic[0].Spare16 := FALSE;
   MH_Hydraulic[1].FLT_Motorprotection := FALSE;
   MH_Hydraulic[1].FLT_Min_Level := FALSE;
   MH_Hydraulic[1].FLT_WRN_C_Max := FALSE;
   MH_Hydraulic[1].FLT_C_Max := FALSE;
   MH_Hydraulic[1].FLT_Filter_HP := FALSE;
   MH_Hydraulic[1].FLT_Filter_backflow := FALSE;
   MH_Hydraulic[1].FLT_cable_break := FALSE;
   MH_Hydraulic[1].FLT_P_Max := FALSE;
   MH_Hydraulic[1].FLT_Moog_Filter := FALSE;
   MH_Hydraulic[1].FLT_MotorProtFilterPump := FALSE;
   MH_Hydraulic[1].FLT_MinLevelFilterPump := FALSE;
   MH_Hydraulic[1].FLT_MaxLevelFilterPump := FALSE;
   MH_Hydraulic[1].FLT_FilterBypass := FALSE;
   MH_Hydraulic[1].Spare14 := FALSE;
   MH_Hydraulic[1].Spare15 := FALSE;
   MH_Hydraulic[1].Spare16 := FALSE;
   MH_Hydraulic[2].FLT_Motorprotection := FALSE;
   MH_Hydraulic[2].FLT_Min_Level := FALSE;
   MH_Hydraulic[2].FLT_WRN_C_Max := FALSE;
   MH_Hydraulic[2].FLT_C_Max := FALSE;
   MH_Hydraulic[2].FLT_Filter_HP := FALSE;
   MH_Hydraulic[2].FLT_Filter_backflow := FALSE;
   MH_Hydraulic[2].FLT_cable_break := FALSE;
   MH_Hydraulic[2].FLT_P_Max := FALSE;
   MH_Hydraulic[2].FLT_Moog_Filter := FALSE;
   MH_Hydraulic[2].FLT_MotorProtFilterPump := FALSE;
   MH_Hydraulic[2].FLT_MinLevelFilterPump := FALSE;
   MH_Hydraulic[2].FLT_MaxLevelFilterPump := FALSE;
   MH_Hydraulic[2].FLT_FilterBypass := FALSE;
   MH_Hydraulic[2].Spare14 := FALSE;
   MH_Hydraulic[2].Spare15 := FALSE;
   MH_Hydraulic[2].Spare16 := FALSE;
   S_Hydraulic[0].FLT_Motorprotection := FALSE;
   S_Hydraulic[0].FLT_Min_Level := FALSE;
   S_Hydraulic[0].FLT_WRN_C_Max := FALSE;
   S_Hydraulic[0].FLT_C_Max := FALSE;
   S_Hydraulic[0].FLT_Filter_HP := FALSE;
   S_Hydraulic[0].FLT_Filter_backflow := FALSE;
   S_Hydraulic[0].FLT_cable_break := FALSE;
   S_Hydraulic[0].FLT_P_Max := FALSE;
   S_Hydraulic[0].FLT_Moog_Filter := FALSE;
   S_Hydraulic[0].FLT_MotorProtFilterPump := FALSE;
   S_Hydraulic[0].FLT_MinLevelFilterPump := FALSE;
   S_Hydraulic[0].FLT_MaxLevelFilterPump := FALSE;
   S_Hydraulic[0].FLT_FilterBypass := FALSE;
   S_Hydraulic[0].Spare14 := FALSE;
   S_Hydraulic[0].Spare15 := FALSE;
   S_Hydraulic[0].Spare16 := FALSE;
   S_Hydraulic[1].FLT_Motorprotection := FALSE;
   S_Hydraulic[1].FLT_Min_Level := FALSE;
   S_Hydraulic[1].FLT_WRN_C_Max := FALSE;
   S_Hydraulic[1].FLT_C_Max := FALSE;
   S_Hydraulic[1].FLT_Filter_HP := FALSE;
   S_Hydraulic[1].FLT_Filter_backflow := FALSE;
   S_Hydraulic[1].FLT_cable_break := FALSE;
   S_Hydraulic[1].FLT_P_Max := FALSE;
   S_Hydraulic[1].FLT_Moog_Filter := FALSE;
   S_Hydraulic[1].FLT_MotorProtFilterPump := FALSE;
   S_Hydraulic[1].FLT_MinLevelFilterPump := FALSE;
   S_Hydraulic[1].FLT_MaxLevelFilterPump := FALSE;
   S_Hydraulic[1].FLT_FilterBypass := FALSE;
   S_Hydraulic[1].Spare14 := FALSE;
   S_Hydraulic[1].Spare15 := FALSE;
   S_Hydraulic[1].Spare16 := FALSE;
   S_Hydraulic[2].FLT_Motorprotection := FALSE;
   S_Hydraulic[2].FLT_Min_Level := FALSE;
   S_Hydraulic[2].FLT_WRN_C_Max := FALSE;
   S_Hydraulic[2].FLT_C_Max := FALSE;
   S_Hydraulic[2].FLT_Filter_HP := FALSE;
   S_Hydraulic[2].FLT_Filter_backflow := FALSE;
   S_Hydraulic[2].FLT_cable_break := FALSE;
   S_Hydraulic[2].FLT_P_Max := FALSE;
   S_Hydraulic[2].FLT_Moog_Filter := FALSE;
   S_Hydraulic[2].FLT_MotorProtFilterPump := FALSE;
   S_Hydraulic[2].FLT_MinLevelFilterPump := FALSE;
   S_Hydraulic[2].FLT_MaxLevelFilterPump := FALSE;
   S_Hydraulic[2].FLT_FilterBypass := FALSE;
   S_Hydraulic[2].Spare14 := FALSE;
   S_Hydraulic[2].Spare15 := FALSE;
   S_Hydraulic[2].Spare16 := FALSE;
   NZL_Hydraulic[0].FLT_Motorprotection := FALSE;
   NZL_Hydraulic[0].FLT_Min_Level := FALSE;
   NZL_Hydraulic[0].FLT_WRN_C_Max := FALSE;
   NZL_Hydraulic[0].FLT_C_Max := FALSE;
   NZL_Hydraulic[0].FLT_Filter_HP := FALSE;
   NZL_Hydraulic[0].FLT_Filter_backflow := FALSE;
   NZL_Hydraulic[0].FLT_cable_break := FALSE;
   NZL_Hydraulic[0].FLT_P_Max := FALSE;
   NZL_Hydraulic[0].FLT_Moog_Filter := FALSE;
   NZL_Hydraulic[0].FLT_MotorProtFilterPump := FALSE;
   NZL_Hydraulic[0].FLT_MinLevelFilterPump := FALSE;
   NZL_Hydraulic[0].FLT_MaxLevelFilterPump := FALSE;
   NZL_Hydraulic[0].FLT_FilterBypass := FALSE;
   NZL_Hydraulic[0].Spare14 := FALSE;
   NZL_Hydraulic[0].Spare15 := FALSE;
   NZL_Hydraulic[0].Spare16 := FALSE;
   NZL_Hydraulic[1].FLT_Motorprotection := FALSE;
   NZL_Hydraulic[1].FLT_Min_Level := FALSE;
   NZL_Hydraulic[1].FLT_WRN_C_Max := FALSE;
   NZL_Hydraulic[1].FLT_C_Max := FALSE;
   NZL_Hydraulic[1].FLT_Filter_HP := FALSE;
   NZL_Hydraulic[1].FLT_Filter_backflow := FALSE;
   NZL_Hydraulic[1].FLT_cable_break := FALSE;
   NZL_Hydraulic[1].FLT_P_Max := FALSE;
   NZL_Hydraulic[1].FLT_Moog_Filter := FALSE;
   NZL_Hydraulic[1].FLT_MotorProtFilterPump := FALSE;
   NZL_Hydraulic[1].FLT_MinLevelFilterPump := FALSE;
   NZL_Hydraulic[1].FLT_MaxLevelFilterPump := FALSE;
   NZL_Hydraulic[1].FLT_FilterBypass := FALSE;
   NZL_Hydraulic[1].Spare14 := FALSE;
   NZL_Hydraulic[1].Spare15 := FALSE;
   NZL_Hydraulic[1].Spare16 := FALSE;
   NZL_Hydraulic[2].FLT_Motorprotection := FALSE;
   NZL_Hydraulic[2].FLT_Min_Level := FALSE;
   NZL_Hydraulic[2].FLT_WRN_C_Max := FALSE;
   NZL_Hydraulic[2].FLT_C_Max := FALSE;
   NZL_Hydraulic[2].FLT_Filter_HP := FALSE;
   NZL_Hydraulic[2].FLT_Filter_backflow := FALSE;
   NZL_Hydraulic[2].FLT_cable_break := FALSE;
   NZL_Hydraulic[2].FLT_P_Max := FALSE;
   NZL_Hydraulic[2].FLT_Moog_Filter := FALSE;
   NZL_Hydraulic[2].FLT_MotorProtFilterPump := FALSE;
   NZL_Hydraulic[2].FLT_MinLevelFilterPump := FALSE;
   NZL_Hydraulic[2].FLT_MaxLevelFilterPump := FALSE;
   NZL_Hydraulic[2].FLT_FilterBypass := FALSE;
   NZL_Hydraulic[2].Spare14 := FALSE;
   NZL_Hydraulic[2].Spare15 := FALSE;
   NZL_Hydraulic[2].Spare16 := FALSE;
   EmergencyStop_Hydraulic[1] := FALSE;
   EmergencyStop_Hydraulic[2] := FALSE;
   EmergencyStop_Hydraulic[3] := FALSE;
   EmergencyStop_Hydraulic[4] := FALSE;
   EmergencyStop_Hydraulic[5] := FALSE;
   EmergencyStop_Hydraulic[6] := FALSE;
   EmergencyStop_Hydraulic[7] := FALSE;
   EmergencyStop_Hydraulic[8] := FALSE;
   EmergencyStop_Hydraulic[9] := FALSE;
   EmergencyStop_Hydraulic[10] := FALSE;
   EmergencyStop_Hydraulic[11] := FALSE;
   EmergencyStop_Hydraulic[12] := FALSE;
   EmergencyStop_Hydraulic[13] := FALSE;
   EmergencyStop_Hydraulic[14] := FALSE;
   EmergencyStop_Hydraulic[15] := FALSE;
   EmergencyStop_Hydraulic[16] := FALSE;
END_DATA_BLOCK

DATA_BLOCK "DB822_Error_Tank"   // DB822
TITLE = Faults general at plant and machine
{ S7_Optimized_Access := 'FALSE' }
VERSION : 0.1
   VAR
      FeedPump : Array[0..12] of "UDT1801_FLT_auxDrive";
      Agitator : Array[0..12] of "UDT1801_Agitator";
      Refilling_Tank : Array[0..12] of "UDT1802_FLT_Tank_Refill";   // Tank, refiling component 1 - 16
      CirculationPump : Array[0..12] of "UDT1801_FLT_auxDrive";
      RefillingStation : Array[0..12] of "UDT1803_FLT_RefilStation";
      Temperature_Heatexchange : Array[0..12] of "UDT1820_FLT_ProcessValue";   // Process value tempering heat exchanger
      ControllerTankTemp : Array[0..12] of "UDT1804_FLT_Controller";   // Controller units
      ControllerTankJacketHeater : Array[0..12] of "UDT1804_FLT_Controller";   // Controller units
      ControllerBarellTemp : Array[0..12] of "UDT1804_FLT_Controller";   // Controller units
      Vacuum : Array[0..12] of "UDT1806_FLT_Vacuum";   // Fault vacuum unit daytank (Level 3)
      CoverLift : Array[0..12] of "UDT1809_FLT_CoverLift";   // Fault cover lift
      LevelRefillingStation : Array[0..12] of "UDT1820_FLT_ProcessValue";   // Process value level refilling station
      TempRefillingStation : Array[0..12] of "UDT1820_FLT_ProcessValue";   // Process value temperature refilling station
      JacketHeater_Tank : Array[0..12] of "UDT1820_FLT_ProcessValue";   // Process value Pressure tank
      LeakageMonitor : Array[0..12] of "UDT1826_FLT_LeakageMonit";   // Leakagemonitor components
      AgitatorBarrel : Array[0..12] of "UDT1801_FLT_auxDrive";
      Pentan : Array[0..12] of "UDT1810_Pentan";
      InterfaceContainer : Struct
         FLT_SupplyContainerstation : Bool;
         FLT_containerstation : Bool;   // Signal container fault existing
         MSG_EScontainerstation : Bool;
         Spare_04 : Bool;
         FLT_containerNotReady_C1 : Bool;
         FLT_containerNotReady_C2 : Bool;
         FLT_containerNotReady_C3 : Bool;
         FLT_containerNotReady_C4 : Bool;
         MSG_containerNotReady_C1 : Bool;
         MSG_containerNotReady_C2 : Bool;
         MSG_containerNotReady_C3 : Bool;
         MSG_containerNotReady_C4 : Bool;
         Spare_13 : Bool;
         Spare_14 : Bool;
         Spare_15 : Bool;
         Spare_16 : Bool;
      END_STRUCT;
   END_VAR
BEGIN
   FeedPump[0].FLT_Motorprotection := FALSE;
   FeedPump[0].FLT_FrequencyConverter := FALSE;
   FeedPump[0].FLT_MaxP_MaxLTripTray := FALSE;
   FeedPump[0].FLT_Dryrunsafety := FALSE;
   FeedPump[0].FLT_wrong_Timevalue := FALSE;
   FeedPump[0].FLT_MaxPressureDiff := FALSE;
   FeedPump[0].Mes_Min_temp := FALSE;
   FeedPump[0].FLT_MotorFan := FALSE;
   FeedPump[0].Mes_Min_Level := FALSE;
   FeedPump[0].FLT_No_Barrel := FALSE;
   FeedPump[0].Mes_No_Barrel := FALSE;
   FeedPump[0].Spare_1_3 := FALSE;
   FeedPump[0].Spare_1_4 := FALSE;
   FeedPump[0].Spare_1_5 := FALSE;
   FeedPump[0].Spare_1_6 := FALSE;
   FeedPump[0].Spare_1_7 := FALSE;
   FeedPump[1].FLT_Motorprotection := FALSE;
   FeedPump[1].FLT_FrequencyConverter := FALSE;
   FeedPump[1].FLT_MaxP_MaxLTripTray := FALSE;
   FeedPump[1].FLT_Dryrunsafety := FALSE;
   FeedPump[1].FLT_wrong_Timevalue := FALSE;
   FeedPump[1].FLT_MaxPressureDiff := FALSE;
   FeedPump[1].Mes_Min_temp := FALSE;
   FeedPump[1].FLT_MotorFan := FALSE;
   FeedPump[1].Mes_Min_Level := FALSE;
   FeedPump[1].FLT_No_Barrel := FALSE;
   FeedPump[1].Mes_No_Barrel := FALSE;
   FeedPump[1].Spare_1_3 := FALSE;
   FeedPump[1].Spare_1_4 := FALSE;
   FeedPump[1].Spare_1_5 := FALSE;
   FeedPump[1].Spare_1_6 := FALSE;
   FeedPump[1].Spare_1_7 := FALSE;
   FeedPump[2].FLT_Motorprotection := FALSE;
   FeedPump[2].FLT_FrequencyConverter := FALSE;
   FeedPump[2].FLT_MaxP_MaxLTripTray := FALSE;
   FeedPump[2].FLT_Dryrunsafety := FALSE;
   FeedPump[2].FLT_wrong_Timevalue := FALSE;
   FeedPump[2].FLT_MaxPressureDiff := FALSE;
   FeedPump[2].Mes_Min_temp := FALSE;
   FeedPump[2].FLT_MotorFan := FALSE;
   FeedPump[2].Mes_Min_Level := FALSE;
   FeedPump[2].FLT_No_Barrel := FALSE;
   FeedPump[2].Mes_No_Barrel := FALSE;
   FeedPump[2].Spare_1_3 := FALSE;
   FeedPump[2].Spare_1_4 := FALSE;
   FeedPump[2].Spare_1_5 := FALSE;
   FeedPump[2].Spare_1_6 := FALSE;
   FeedPump[2].Spare_1_7 := FALSE;
   FeedPump[3].FLT_Motorprotection := FALSE;
   FeedPump[3].FLT_FrequencyConverter := FALSE;
   FeedPump[3].FLT_MaxP_MaxLTripTray := FALSE;
   FeedPump[3].FLT_Dryrunsafety := FALSE;
   FeedPump[3].FLT_wrong_Timevalue := FALSE;
   FeedPump[3].FLT_MaxPressureDiff := FALSE;
   FeedPump[3].Mes_Min_temp := FALSE;
   FeedPump[3].FLT_MotorFan := FALSE;
   FeedPump[3].Mes_Min_Level := FALSE;
   FeedPump[3].FLT_No_Barrel := FALSE;
   FeedPump[3].Mes_No_Barrel := FALSE;
   FeedPump[3].Spare_1_3 := FALSE;
   FeedPump[3].Spare_1_4 := FALSE;
   FeedPump[3].Spare_1_5 := FALSE;
   FeedPump[3].Spare_1_6 := FALSE;
   FeedPump[3].Spare_1_7 := FALSE;
   FeedPump[4].FLT_Motorprotection := FALSE;
   FeedPump[4].FLT_FrequencyConverter := FALSE;
   FeedPump[4].FLT_MaxP_MaxLTripTray := FALSE;
   FeedPump[4].FLT_Dryrunsafety := FALSE;
   FeedPump[4].FLT_wrong_Timevalue := FALSE;
   FeedPump[4].FLT_MaxPressureDiff := FALSE;
   FeedPump[4].Mes_Min_temp := FALSE;
   FeedPump[4].FLT_MotorFan := FALSE;
   FeedPump[4].Mes_Min_Level := FALSE;
   FeedPump[4].FLT_No_Barrel := FALSE;
   FeedPump[4].Mes_No_Barrel := FALSE;
   FeedPump[4].Spare_1_3 := FALSE;
   FeedPump[4].Spare_1_4 := FALSE;
   FeedPump[4].Spare_1_5 := FALSE;
   FeedPump[4].Spare_1_6 := FALSE;
   FeedPump[4].Spare_1_7 := FALSE;
   FeedPump[5].FLT_Motorprotection := FALSE;
   FeedPump[5].FLT_FrequencyConverter := FALSE;
   FeedPump[5].FLT_MaxP_MaxLTripTray := FALSE;
   FeedPump[5].FLT_Dryrunsafety := FALSE;
   FeedPump[5].FLT_wrong_Timevalue := FALSE;
   FeedPump[5].FLT_MaxPressureDiff := FALSE;
   FeedPump[5].Mes_Min_temp := FALSE;
   FeedPump[5].FLT_MotorFan := FALSE;
   FeedPump[5].Mes_Min_Level := FALSE;
   FeedPump[5].FLT_No_Barrel := FALSE;
   FeedPump[5].Mes_No_Barrel := FALSE;
   FeedPump[5].Spare_1_3 := FALSE;
   FeedPump[5].Spare_1_4 := FALSE;
   FeedPump[5].Spare_1_5 := FALSE;
   FeedPump[5].Spare_1_6 := FALSE;
   FeedPump[5].Spare_1_7 := FALSE;
   FeedPump[6].FLT_Motorprotection := FALSE;
   FeedPump[6].FLT_FrequencyConverter := FALSE;
   FeedPump[6].FLT_MaxP_MaxLTripTray := FALSE;
   FeedPump[6].FLT_Dryrunsafety := FALSE;
   FeedPump[6].FLT_wrong_Timevalue := FALSE;
   FeedPump[6].FLT_MaxPressureDiff := FALSE;
   FeedPump[6].Mes_Min_temp := FALSE;
   FeedPump[6].FLT_MotorFan := FALSE;
   FeedPump[6].Mes_Min_Level := FALSE;
   FeedPump[6].FLT_No_Barrel := FALSE;
   FeedPump[6].Mes_No_Barrel := FALSE;
   FeedPump[6].Spare_1_3 := FALSE;
   FeedPump[6].Spare_1_4 := FALSE;
   FeedPump[6].Spare_1_5 := FALSE;
   FeedPump[6].Spare_1_6 := FALSE;
   FeedPump[6].Spare_1_7 := FALSE;
   FeedPump[7].FLT_Motorprotection := FALSE;
   FeedPump[7].FLT_FrequencyConverter := FALSE;
   FeedPump[7].FLT_MaxP_MaxLTripTray := FALSE;
   FeedPump[7].FLT_Dryrunsafety := FALSE;
   FeedPump[7].FLT_wrong_Timevalue := FALSE;
   FeedPump[7].FLT_MaxPressureDiff := FALSE;
   FeedPump[7].Mes_Min_temp := FALSE;
   FeedPump[7].FLT_MotorFan := FALSE;
   FeedPump[7].Mes_Min_Level := FALSE;
   FeedPump[7].FLT_No_Barrel := FALSE;
   FeedPump[7].Mes_No_Barrel := FALSE;
   FeedPump[7].Spare_1_3 := FALSE;
   FeedPump[7].Spare_1_4 := FALSE;
   FeedPump[7].Spare_1_5 := FALSE;
   FeedPump[7].Spare_1_6 := FALSE;
   FeedPump[7].Spare_1_7 := FALSE;
   FeedPump[8].FLT_Motorprotection := FALSE;
   FeedPump[8].FLT_FrequencyConverter := FALSE;
   FeedPump[8].FLT_MaxP_MaxLTripTray := FALSE;
   FeedPump[8].FLT_Dryrunsafety := FALSE;
   FeedPump[8].FLT_wrong_Timevalue := FALSE;
   FeedPump[8].FLT_MaxPressureDiff := FALSE;
   FeedPump[8].Mes_Min_temp := FALSE;
   FeedPump[8].FLT_MotorFan := FALSE;
   FeedPump[8].Mes_Min_Level := FALSE;
   FeedPump[8].FLT_No_Barrel := FALSE;
   FeedPump[8].Mes_No_Barrel := FALSE;
   FeedPump[8].Spare_1_3 := FALSE;
   FeedPump[8].Spare_1_4 := FALSE;
   FeedPump[8].Spare_1_5 := FALSE;
   FeedPump[8].Spare_1_6 := FALSE;
   FeedPump[8].Spare_1_7 := FALSE;
   FeedPump[9].FLT_Motorprotection := FALSE;
   FeedPump[9].FLT_FrequencyConverter := FALSE;
   FeedPump[9].FLT_MaxP_MaxLTripTray := FALSE;
   FeedPump[9].FLT_Dryrunsafety := FALSE;
   FeedPump[9].FLT_wrong_Timevalue := FALSE;
   FeedPump[9].FLT_MaxPressureDiff := FALSE;
   FeedPump[9].Mes_Min_temp := FALSE;
   FeedPump[9].FLT_MotorFan := FALSE;
   FeedPump[9].Mes_Min_Level := FALSE;
   FeedPump[9].FLT_No_Barrel := FALSE;
   FeedPump[9].Mes_No_Barrel := FALSE;
   FeedPump[9].Spare_1_3 := FALSE;
   FeedPump[9].Spare_1_4 := FALSE;
   FeedPump[9].Spare_1_5 := FALSE;
   FeedPump[9].Spare_1_6 := FALSE;
   FeedPump[9].Spare_1_7 := FALSE;
   FeedPump[10].FLT_Motorprotection := FALSE;
   FeedPump[10].FLT_FrequencyConverter := FALSE;
   FeedPump[10].FLT_MaxP_MaxLTripTray := FALSE;
   FeedPump[10].FLT_Dryrunsafety := FALSE;
   FeedPump[10].FLT_wrong_Timevalue := FALSE;
   FeedPump[10].FLT_MaxPressureDiff := FALSE;
   FeedPump[10].Mes_Min_temp := FALSE;
   FeedPump[10].FLT_MotorFan := FALSE;
   FeedPump[10].Mes_Min_Level := FALSE;
   FeedPump[10].FLT_No_Barrel := FALSE;
   FeedPump[10].Mes_No_Barrel := FALSE;
   FeedPump[10].Spare_1_3 := FALSE;
   FeedPump[10].Spare_1_4 := FALSE;
   FeedPump[10].Spare_1_5 := FALSE;
   FeedPump[10].Spare_1_6 := FALSE;
   FeedPump[10].Spare_1_7 := FALSE;
   FeedPump[11].FLT_Motorprotection := FALSE;
   FeedPump[11].FLT_FrequencyConverter := FALSE;
   FeedPump[11].FLT_MaxP_MaxLTripTray := FALSE;
   FeedPump[11].FLT_Dryrunsafety := FALSE;
   FeedPump[11].FLT_wrong_Timevalue := FALSE;
   FeedPump[11].FLT_MaxPressureDiff := FALSE;
   FeedPump[11].Mes_Min_temp := FALSE;
   FeedPump[11].FLT_MotorFan := FALSE;
   FeedPump[11].Mes_Min_Level := FALSE;
   FeedPump[11].FLT_No_Barrel := FALSE;
   FeedPump[11].Mes_No_Barrel := FALSE;
   FeedPump[11].Spare_1_3 := FALSE;
   FeedPump[11].Spare_1_4 := FALSE;
   FeedPump[11].Spare_1_5 := FALSE;
   FeedPump[11].Spare_1_6 := FALSE;
   FeedPump[11].Spare_1_7 := FALSE;
   FeedPump[12].FLT_Motorprotection := FALSE;
   FeedPump[12].FLT_FrequencyConverter := FALSE;
   FeedPump[12].FLT_MaxP_MaxLTripTray := FALSE;
   FeedPump[12].FLT_Dryrunsafety := FALSE;
   FeedPump[12].FLT_wrong_Timevalue := FALSE;
   FeedPump[12].FLT_MaxPressureDiff := FALSE;
   FeedPump[12].Mes_Min_temp := FALSE;
   FeedPump[12].FLT_MotorFan := FALSE;
   // 3450 more start values not shown
END_DATA_BLOCK

